// TIA Portal project "GzyHzy_1500" (V15) (continued)
DATA_BLOCK "模拟量"   // DB2
{ S7_Optimized_Access := 'FALSE' }
VERSION : 0.1
   VAR
      STAT0 : Int;
      STAT1 : Int;
      STAT2 : Int;
      STAT3 : Int;
      STAT4 : Int;
      STAT5 : Int;
      STAT6 : Int;
      STAT7 : Int;
      STAT8 : Int;
      STAT9 : Real;
      STAT10 : Real;
      STAT11 : Real;
      STAT12 : Real;
      STAT13 : Real;
      STAT14 : Real;
      STAT15 : Real;
      STAT16 : Real;
      STAT17 : Real;
      STAT18 : Real;
      STAT19 : Real;
      STAT20 : Real;
      STAT21 : Real;
      STAT22 : Real;
      STAT23 : Real;
      STAT24 : Real;
      STAT25 : Real;
      STAT26 : Real;
      STAT27 : Real;
      STAT28 : Real;
      STAT29 : Real;
      STAT30 : Real;
      STAT31 : Real;
      STAT32 : Real;
      STAT33 : Real;
      STAT34 : Real;
      STAT35 : Real;
      STAT36 : Real;
      STAT37 : Real;
      STAT38 : Real;
      STAT39 : Real;
      STAT40 : Real;
      STAT41 : Real;
      STAT42 : Real;
      STAT43 : Real;
      STAT44 : Real;
      STAT45 : Real;
      STAT46 : Real;
      STAT47 : Real;
      STAT48 : Real;
      STAT49 : Real;
      STAT50 : Real;
      STAT51 : Real;
      STAT52 : Real;
      STAT53 : Real;
      STAT54 : Real;
      STAT55 : Real;
      STAT56 : Real;
      STAT57 : Real;
      STAT58 : Real;
      STAT59 : Real;
      STAT60 : Real;
      STAT61 : Real;
      STAT62 : Real;
      STAT63 : Real;
      STAT64 : Real;
      STAT65 : Real;
      STAT66 : Real;
      STAT67 : Real;
      STAT68 : Real;
      STAT69 : Real;
      STAT70 : Real;
      STAT71 : Real;
      STAT72 : Real;
      STAT73 : Real;
      STAT74 : Real;
      STAT75 : Real;
      STAT76 : Real;
      STAT77 : Real;
      STAT78 : Real;
      STAT79 : Real;
      STAT80 : Real;
      STAT81 : Real;
   END_VAR
BEGIN
END_DATA_BLOCK

DATA_BLOCK "给煤机班累计DB块"   // DB3
{ S7_Optimized_Access := 'FALSE' }
VERSION : 0.0
// stored: InstanceOfName 累计功能块
"累计功能块"
BEGIN
END_DATA_BLOCK

DATA_BLOCK "给煤机日累计DB块"   // DB4
{ S7_Optimized_Access := 'FALSE' }
VERSION : 0.0
// stored: InstanceOfName 累计功能块
"累计功能块"
BEGIN
END_DATA_BLOCK

DATA_BLOCK "给煤机总累计DB块"   // DB5
{ S7_Optimized_Access := 'FALSE' }
VERSION : 0.0
// stored: InstanceOfName 累计功能块
"累计功能块"
BEGIN
END_DATA_BLOCK

DATA_BLOCK "DB6_皮带秤粘料"   // DB6
{ S7_Optimized_Access := 'FALSE' }
VERSION : 0.1
   VAR
      干燥窑定量给煤机给定反馈差值 : Real;
      干燥窑定量给煤机给定反馈差值绝对值 : Real;
      real3 : Real;
      real4 : Real;
      real5 : Real;
      real6 : Real;
      real7 : Real;
      real8 : Real;
      real9 : Real;
      real10 : Real;
      real11 : Real;
      real12 : Real;
      real13 : Real;
      real14 : Real;
      real15 : Real;
      real16 : Real;
      real17 : Real;
      real18 : Real;
      real19 : Real;
      real20 : Real;
      干燥窑定量给煤机粘料报警 : Bool;
      bool2 : Bool;
      bool3 : Bool;
      bool4 : Bool;
      bool5 : Bool;
      bool6 : Bool;
      bool7 : Bool;
      bool8 : Bool;
      bool9 : Bool;
      bool10 : Bool;
      bool11 : Bool;
      bool12 : Bool;
      bool13 : Bool;
      bool14 : Bool;
      bool15 : Bool;
      bool16 : Bool;
      bool17 : Bool;
      bool18 : Bool;
      bool19 : Bool;
      bool20 : Bool;
      bool21 : Bool;
   END_VAR
BEGIN
END_DATA_BLOCK

DATA_BLOCK "累计功能块2_DB"   // DB7
{ S7_Optimized_Access := 'FALSE' }
VERSION : 0.1
// stored: InstanceOfName 累计功能块2
"累计功能块2"
BEGIN
END_DATA_BLOCK

DATA_BLOCK "通讯仪表数据"   // DB20
{ S7_Optimized_Access := 'FALSE' }
VERSION : 0.1
   VAR
      STAT0 : Int;
      "1#窑A档油温1" : Real := 33.4;
      "1#窑A档油温2" : Real := 33.0;
      "1#窑A档油温3" : Real := 34.3;
      "1#窑A档油温4" : Real := 34.0;
      "1#窑A档轴温1" : Real := 33.6;
      "1#窑A档轴温2" : Real := 33.4;
      "1#窑A档轴温3" : Real := 33.6;
      "1#窑A档轴温4" : Real := 34.5;
      "1#窑B档油温1" : Real := 34.3;
      "1#窑B档油温2" : Real := 34.5;
      "1#窑B档油温3" : Real := 35.0;
      "1#窑B档油温4" : Real := 36.1;
      "1#窑B档轴温1" : Real := 34.9;
      "1#窑B档轴温2" : Real := 36.4;
      "1#窑B档轴温3" : Real := 34.9;
      "1#窑B档轴温4" : Real := 36.2;
      "1#窑主电机A相绕组温度" : Real := 62.7;
      "1#窑主电机B相绕组温度" : Real := 63.4;
      "1#窑主电机C相绕组温度" : Real := 62.0;
      "1#窑主电机前轴承温度" : Real := 45.0;
      "1#窑主电机后轴承温度" : Real := 41.8;
      STAT22 : Real;
      STAT23 : Real;
      STAT24 : Real;
      STAT25 : Real;
      STAT26 : Real;
      STAT27 : Real;
      STAT28 : Real;
      STAT29 : Real;
      STAT30 : Real;
      STAT31 : Real;
      STAT32 : Real;
      "1#干燥窑煤粉仓称重" : Real := 11.52;   // 1#干燥窑煤粉仓称重
      STAT34 : Real;
   END_VAR
BEGIN
END_DATA_BLOCK

DATA_BLOCK "模拟量数据"   // DB21
{ S7_Optimized_Access := 'FALSE' }
VERSION : 0.1
   VAR
      "1#干燥窑主电机转速" : Real := 795.8328;
      "1#干燥窑主电机电流" : Real := 246.3866;
      STAT2 : Real;
      "1#干燥窑一次风机运行电流" : Real := 48.19213;
      "1#二次风机运行频率" : Real := 29.89005;
      "1#二次风机运行电流" : Real := 89.02026;
      "1#干燥窑窑尾烟气管道压力" : Real := -16.14584;
      "1#备用一次风机运行电流" : Real := 48.94907;
      "1#备用二次风机运行频率" : Real := 0.1157407;
      "1#备用二次风机运行电流" : Real;
      "1#干燥窑煤粉流量" : Real := 2.039641;
      "1#干燥窑进口烟气管道压力" : Real := -66.84027;
      "1#干燥窑一次风机压力" : Real := 2421.875;
      "1#干燥窑二次风机压力" : Real := 1265.625;
      "1#干燥窑煤粉仓压力" : Real := 11.63208;
      "1#干燥窑燃烧室压力" : Real := -751.3021;
      "1#干燥窑煤粉仓温度1" : Real := 17.85301;
      "1#干燥窑煤粉仓温度2" : Real := 35.30093;
      "1#干燥窑煤粉仓温度3" : Real := 33.96991;
      "1#干燥窑煤粉仓温度4" : Real := 35.3588;
      "1#干燥窑窑尾罩温度" : Real := 194.8495;
      "1#干燥窑进口烟气管道温度" : Real := 346.0648;
      "1#干燥窑燃烧室温度" : Real := 883.3333;
      "1#干燥窑混合室温度" : Real := 426.1863;
      "1#干燥窑主机转速给定" : Real := 800.0;
      "1#干燥窑煤粉仓流量给定" : Real := 2.0;
      振动筛转速给定 : Real;
      STAT27 : Real;
      STAT28 : Real;
      "1#二次风机频率给定" : Real := 30.0;
      STAT30 : Real;
      "1#备用二次风机频率给定" : Real := 38.0;
      "1#干燥窑定量给煤机班累计" : Real := 0.004813849;
      "1#干燥窑定量给煤机日累计" : Real := 362.4617;
      "1#干燥窑定量给煤机总累计" : Real := 362.4611;
      STAT35 : Real;
      STAT36 : Real;
      振动筛转速 : Real;
      振动筛电流 : Real;
   END_VAR
BEGIN
END_DATA_BLOCK

DATA_BLOCK "窑联锁"   // DB23
{ S7_Optimized_Access := 'FALSE' }
VERSION : 0.1
   VAR
      STAT0 : Bool := TRUE;
      STAT1 : Bool;
      STAT2 : Bool;
      STAT3 : Bool;
      STAT4 : Bool;
      STAT5 : Bool;
      STAT6 : Bool;
      STAT7 : Bool;
      STAT8 : Bool := TRUE;
      STAT9 : Bool;
      STAT10 : Bool;
      STAT11 : Bool;
      STAT12 : Bool;
      STAT13 : Bool;
      STAT14 : Bool;
      STAT15 : Bool;
      STAT16 : Bool;
      STAT17 : Bool;
      STAT18 : Word;
   END_VAR
BEGIN
END_DATA_BLOCK

DATA_BLOCK "DB26"   // DB26
{ S7_Optimized_Access := 'FALSE' }
VERSION : 0.1
   VAR
      STAT0 : Bool;
      STAT1 : Bool;
      STAT2 : Bool;
      STAT3 : Bool;
      STAT4 : Bool;
      STAT5 : Bool;
      STAT6 : Bool;
      STAT7 : Bool;
      STAT8 : Word := WORD#16#0002;
      STAT9 : Word;
      STAT10 : Word;
   END_VAR
BEGIN
END_DATA_BLOCK

DATA_BLOCK "FB40_DATA_ALARM_DB"   // DB40
{ S7_Optimized_Access := 'FALSE' }
VERSION : 0.1
// stored: InstanceOfName FB40_DATA_ALARM
"FB40_DATA_ALARM"
BEGIN
END_DATA_BLOCK

FUNCTION_BLOCK "累计功能块"   // FB10, STL
{ S7_Optimized_Access := 'FALSE' }
VERSION : 0.1
   VAR_INPUT
      IN0 : Real;
      IN1 : Bool;
   END_VAR
   VAR_OUTPUT
      OUT2 : Real;
   END_VAR
   VAR
      STAT3 : Real;
      STAT4 : Real;
      STAT5 : Real;
   END_VAR
BEGIN

REGION Network 1
         A(;
         A(;
         A(;
         L     #IN0;
         L     3600.0;
         /R;
         T     #STAT3;
         AN    OV;
         SAVE;
         CLR;
         A     BR;
         );
         JNB   M001;
         L     #STAT3;
         L     10.0;
         /R;
         T     #STAT4;
         AN    OV;
         SAVE;
         CLR;
   M001: A     BR;
         );
         JNB   M002;
         L     #STAT4;
         L     #STAT5;
         +R;
         T     #STAT5;
         AN    OV;
         SAVE;
         CLR;
   M002: A     BR;
         );
         JNB   M003;
         L     #STAT5;
         T     #OUT2;
   M003: NOP   0;
END_REGION

REGION Network 2
         A     #IN1;
         =     %L0.0;
         A     %L0.0;
         JNB   M004;
         L     0.0;
         T     #STAT3;
   M004: NOP   0;
         A     %L0.0;
         JNB   M005;
         L     0.0;
         T     #STAT4;
   M005: NOP   0;
         A     %L0.0;
         JNB   M006;
         L     0.0;
         T     #STAT5;
   M006: NOP   0;
END_REGION

REGION Network 3
         SET;
         SAVE;
END_REGION
END_FUNCTION_BLOCK

FUNCTION_BLOCK "FB40_DATA_ALARM"   // FB40, LAD
{ S7_Optimized_Access := 'FALSE' }
VERSION : 0.1
   VAR
      "1#干燥窑主传动转速" : "FB330_DATA_ALARM";
      "1#干燥窑主传动电流" : "FB330_DATA_ALARM";
      "1#干燥窑二次风机电流" : "FB330_DATA_ALARM";
      "1#干燥窑一次风机电流" : "FB330_DATA_ALARM";
      "1#干燥窑二次风机频率" : "FB330_DATA_ALARM";
      "1#干燥窑窑尾压力" : "FB330_DATA_ALARM";
      "1#干燥窑备用一次风机频率" : "FB330_DATA_ALARM";
      "1#干燥窑备用一次风机电流" : "FB330_DATA_ALARM";
      "1#干燥窑备用二次风机频率" : "FB330_DATA_ALARM";
      "1#干燥窑备用二次风机电流" : "FB330_DATA_ALARM";
      定量给煤机流量 : "FB330_DATA_ALARM";
      烟气管道进口压力 : "FB330_DATA_ALARM";
      "1#干燥窑一次风压" : "FB330_DATA_ALARM";
      "1#干燥窑二次风压" : "FB330_DATA_ALARM";
      煤粉仓压力 : "FB330_DATA_ALARM";
      混合室压力 : "FB330_DATA_ALARM";
      "煤粉仓温度1(PT100)" : "FB330_DATA_ALARM";
      "煤粉仓温度2(PT100)" : "FB330_DATA_ALARM";
      "煤粉仓温度3(PT100)" : "FB330_DATA_ALARM";
      "煤粉仓温度4(PT100)" : "FB330_DATA_ALARM";
      "窑尾温度 K偶" : "FB330_DATA_ALARM";
      "烟气管道进口温度 K偶" : "FB330_DATA_ALARM";
      "燃烧室温度 4~20mA" : "FB330_DATA_ALARM";
      "混合室温度 4~20mA" : "FB330_DATA_ALARM";
      "1#干燥窑进料口压力" : "FB330_DATA_ALARM";
      "1#给煤机出料口负压" : "FB330_DATA_ALARM";
      振动筛转速 : "FB330_DATA_ALARM";
      振动筛电流 : "FB330_DATA_ALARM";
      PIW312 : "FB330_DATA_ALARM";
      PIW314 : "FB330_DATA_ALARM";
      PIW316 : "FB330_DATA_ALARM";
      PIW318 : "FB330_DATA_ALARM";
      "1#窑A档轴温1" : "FB330_DATA_ALARM";
      "1#窑A档油温1" : "FB330_DATA_ALARM";
      "1#窑A档轴温2" : "FB330_DATA_ALARM";
      "1#窑A档油温2" : "FB330_DATA_ALARM";
      "1#窑A档轴温3" : "FB330_DATA_ALARM";
      "1#窑A档油温3" : "FB330_DATA_ALARM";
      "1#窑A档轴温4" : "FB330_DATA_ALARM";
      "1#窑A档油温4" : "FB330_DATA_ALARM";
      "1#窑B档轴温1" : "FB330_DATA_ALARM";
      "1#窑B档油温1" : "FB330_DATA_ALARM";
      "1#窑B档轴温2" : "FB330_DATA_ALARM";
      "1#窑B档油温2" : "FB330_DATA_ALARM";
      "1#窑B档轴温3" : "FB330_DATA_ALARM";
      "1#窑B档油温3" : "FB330_DATA_ALARM";
      "1#窑B档轴温4" : "FB330_DATA_ALARM";
      "1#窑B档油温4" : "FB330_DATA_ALARM";
      "1#窑主电机A相绕组温度" : "FB330_DATA_ALARM";
      "1#窑主电机B相绕组温度" : "FB330_DATA_ALARM";
      "1#窑主电机C相绕组温度" : "FB330_DATA_ALARM";
      "1#窑主电机前轴承温度" : "FB330_DATA_ALARM";
      "1#窑主电机后轴承温度" : "FB330_DATA_ALARM";
      PID404 : "FB330_DATA_ALARM";
      PID408 : "FB330_DATA_ALARM";
      PID412 : "FB330_DATA_ALARM";
      "1#干燥窑煤粉仓称重" : "FB330_DATA_ALARM";
      STATIC1 : "FB330_DATA_ALARM";
      STATIC2 : "FB330_DATA_ALARM";
      STATIC3 : "FB330_DATA_ALARM";
   END_VAR
   VAR_TEMP
      TEMP1 : Real;
   END_VAR
BEGIN

REGION Network 1
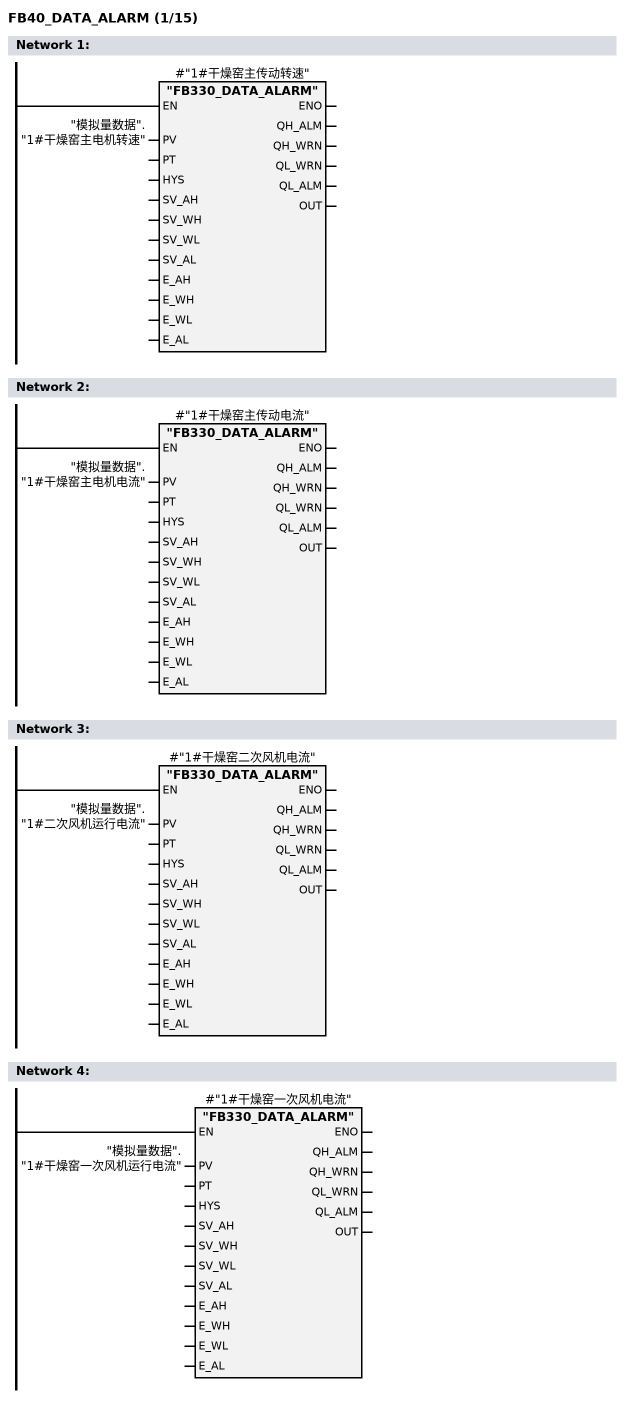
   RUNG wire#powerrail
      #"1#干燥窑主传动转速"(PV := "模拟量数据"."1#干燥窑主电机转速", PT :=, HYS :=, SV_AH :=, SV_WH :=, SV_WL :=, SV_AL :=, E_AH :=, E_WH :=, E_WL :=, E_AL :=, QH_ALM =>, QH_WRN =>, QL_WRN =>, QL_ALM =>, OUT =>)
   END_RUNG
   // the same network as SCL:
   #"1#干燥窑主传动转速"(PV := "模拟量数据"."1#干燥窑主电机转速");   // "FB330_DATA_ALARM"
END_REGION

REGION Network 2
   RUNG wire#powerrail
      #"1#干燥窑主传动电流"(PV := "模拟量数据"."1#干燥窑主电机电流", PT :=, HYS :=, SV_AH :=, SV_WH :=, SV_WL :=, SV_AL :=, E_AH :=, E_WH :=, E_WL :=, E_AL :=, QH_ALM =>, QH_WRN =>, QL_WRN =>, QL_ALM =>, OUT =>)
   END_RUNG
   // the same network as SCL:
   #"1#干燥窑主传动电流"(PV := "模拟量数据"."1#干燥窑主电机电流");   // "FB330_DATA_ALARM"
END_REGION

REGION Network 3
   RUNG wire#powerrail
      #"1#干燥窑二次风机电流"(PV := "模拟量数据"."1#二次风机运行电流", PT :=, HYS :=, SV_AH :=, SV_WH :=, SV_WL :=, SV_AL :=, E_AH :=, E_WH :=, E_WL :=, E_AL :=, QH_ALM =>, QH_WRN =>, QL_WRN =>, QL_ALM =>, OUT =>)
   END_RUNG
   // the same network as SCL:
   #"1#干燥窑二次风机电流"(PV := "模拟量数据"."1#二次风机运行电流");   // "FB330_DATA_ALARM"
END_REGION

REGION Network 4
   RUNG wire#powerrail
      #"1#干燥窑一次风机电流"(PV := "模拟量数据"."1#干燥窑一次风机运行电流", PT :=, HYS :=, SV_AH :=, SV_WH :=, SV_WL :=, SV_AL :=, E_AH :=, E_WH :=, E_WL :=, E_AL :=, QH_ALM =>, QH_WRN =>, QL_WRN =>, QL_ALM =>, OUT =>)
   END_RUNG
   // the same network as SCL:
   #"1#干燥窑一次风机电流"(PV := "模拟量数据"."1#干燥窑一次风机运行电流");   // "FB330_DATA_ALARM"
END_REGION

REGION Network 5
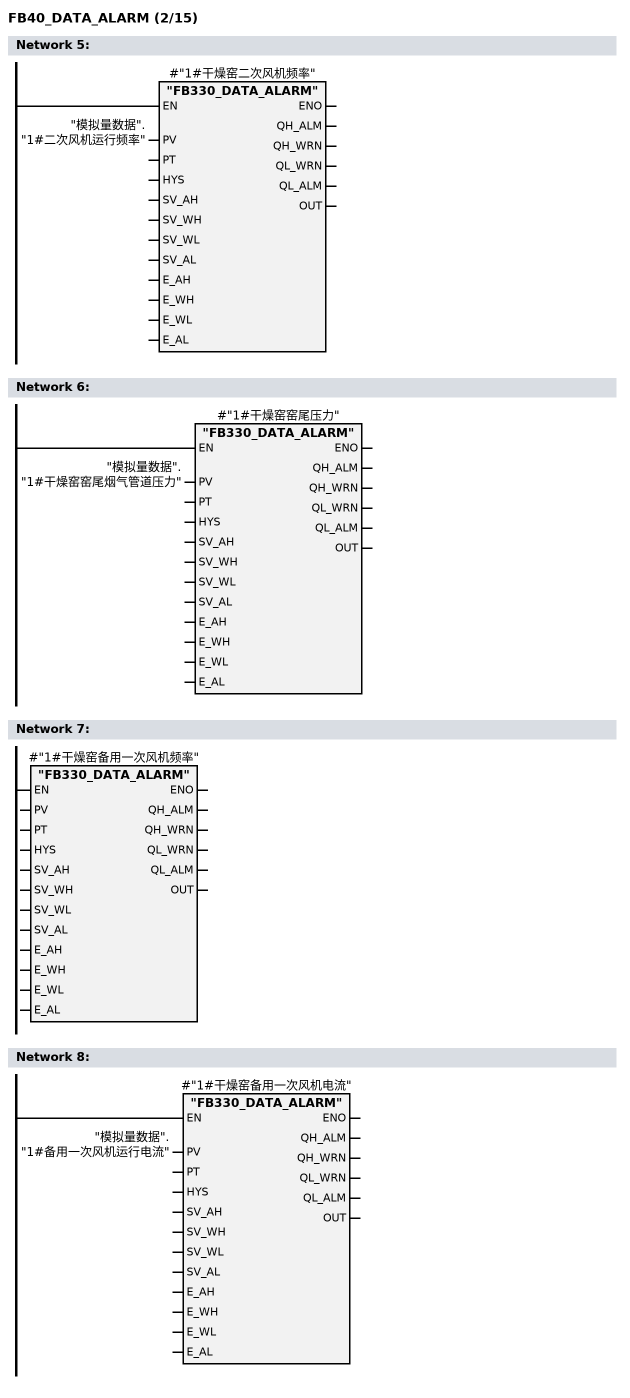
   RUNG wire#powerrail
      #"1#干燥窑二次风机频率"(PV := "模拟量数据"."1#二次风机运行频率", PT :=, HYS :=, SV_AH :=, SV_WH :=, SV_WL :=, SV_AL :=, E_AH :=, E_WH :=, E_WL :=, E_AL :=, QH_ALM =>, QH_WRN =>, QL_WRN =>, QL_ALM =>, OUT =>)
   END_RUNG
   // the same network as SCL:
   #"1#干燥窑二次风机频率"(PV := "模拟量数据"."1#二次风机运行频率");   // "FB330_DATA_ALARM"
END_REGION

REGION Network 6
   RUNG wire#powerrail
      #"1#干燥窑窑尾压力"(PV := "模拟量数据"."1#干燥窑窑尾烟气管道压力", PT :=, HYS :=, SV_AH :=, SV_WH :=, SV_WL :=, SV_AL :=, E_AH :=, E_WH :=, E_WL :=, E_AL :=, QH_ALM =>, QH_WRN =>, QL_WRN =>, QL_ALM =>, OUT =>)
   END_RUNG
   // the same network as SCL:
   #"1#干燥窑窑尾压力"(PV := "模拟量数据"."1#干燥窑窑尾烟气管道压力");   // "FB330_DATA_ALARM"
END_REGION

REGION Network 7
   RUNG wire#powerrail
      #"1#干燥窑备用一次风机频率"(PV :=, PT :=, HYS :=, SV_AH :=, SV_WH :=, SV_WL :=, SV_AL :=, E_AH :=, E_WH :=, E_WL :=, E_AL :=, QH_ALM =>, QH_WRN =>, QL_WRN =>, QL_ALM =>, OUT =>)
   END_RUNG
   // the same network as SCL:
   #"1#干燥窑备用一次风机频率"();   // "FB330_DATA_ALARM"
END_REGION

REGION Network 8
   RUNG wire#powerrail
      #"1#干燥窑备用一次风机电流"(PV := "模拟量数据"."1#备用一次风机运行电流", PT :=, HYS :=, SV_AH :=, SV_WH :=, SV_WL :=, SV_AL :=, E_AH :=, E_WH :=, E_WL :=, E_AL :=, QH_ALM =>, QH_WRN =>, QL_WRN =>, QL_ALM =>, OUT =>)
   END_RUNG
   // the same network as SCL:
   #"1#干燥窑备用一次风机电流"(PV := "模拟量数据"."1#备用一次风机运行电流");   // "FB330_DATA_ALARM"
END_REGION

REGION Network 9
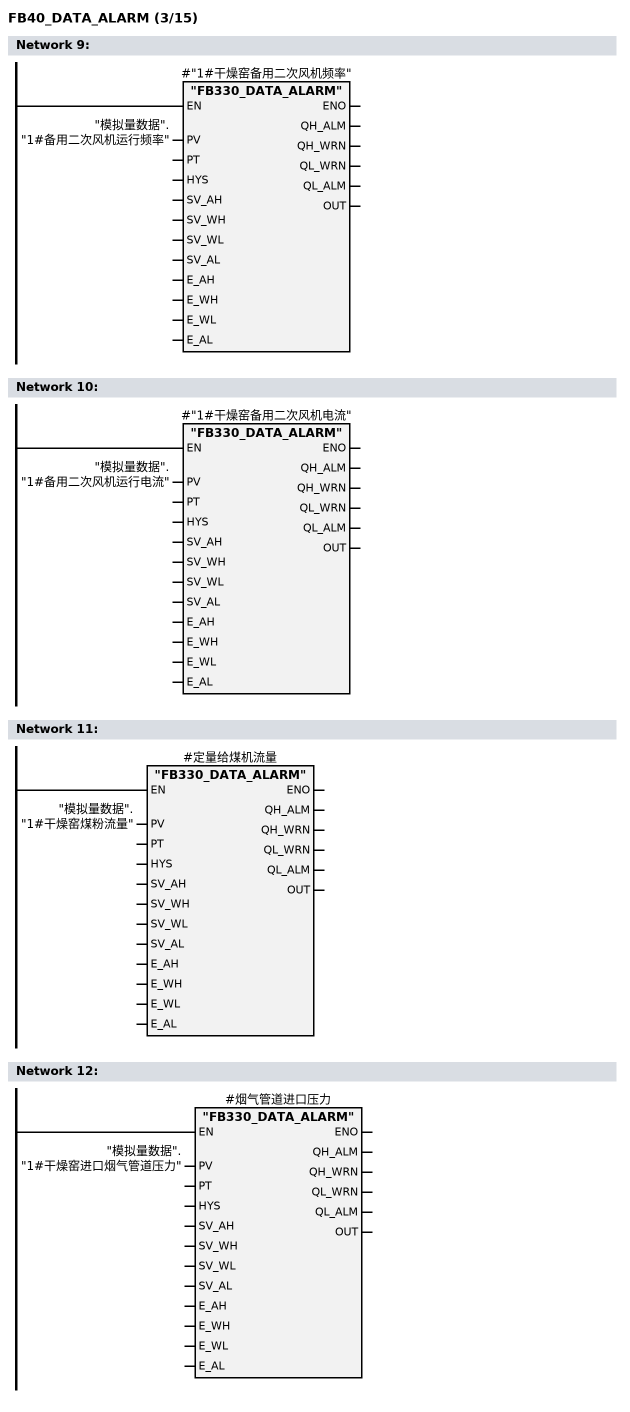
   RUNG wire#powerrail
      #"1#干燥窑备用二次风机频率"(PV := "模拟量数据"."1#备用二次风机运行频率", PT :=, HYS :=, SV_AH :=, SV_WH :=, SV_WL :=, SV_AL :=, E_AH :=, E_WH :=, E_WL :=, E_AL :=, QH_ALM =>, QH_WRN =>, QL_WRN =>, QL_ALM =>, OUT =>)
   END_RUNG
   // the same network as SCL:
   #"1#干燥窑备用二次风机频率"(PV := "模拟量数据"."1#备用二次风机运行频率");   // "FB330_DATA_ALARM"
END_REGION

REGION Network 10
   RUNG wire#powerrail
      #"1#干燥窑备用二次风机电流"(PV := "模拟量数据"."1#备用二次风机运行电流", PT :=, HYS :=, SV_AH :=, SV_WH :=, SV_WL :=, SV_AL :=, E_AH :=, E_WH :=, E_WL :=, E_AL :=, QH_ALM =>, QH_WRN =>, QL_WRN =>, QL_ALM =>, OUT =>)
   END_RUNG
   // the same network as SCL:
   #"1#干燥窑备用二次风机电流"(PV := "模拟量数据"."1#备用二次风机运行电流");   // "FB330_DATA_ALARM"
END_REGION

REGION Network 11
   RUNG wire#powerrail
      #定量给煤机流量(PV := "模拟量数据"."1#干燥窑煤粉流量", PT :=, HYS :=, SV_AH :=, SV_WH :=, SV_WL :=, SV_AL :=, E_AH :=, E_WH :=, E_WL :=, E_AL :=, QH_ALM =>, QH_WRN =>, QL_WRN =>, QL_ALM =>, OUT =>)
   END_RUNG
   // the same network as SCL:
   #定量给煤机流量(PV := "模拟量数据"."1#干燥窑煤粉流量");   // "FB330_DATA_ALARM"
END_REGION

REGION Network 12
   RUNG wire#powerrail
      #烟气管道进口压力(PV := "模拟量数据"."1#干燥窑进口烟气管道压力", PT :=, HYS :=, SV_AH :=, SV_WH :=, SV_WL :=, SV_AL :=, E_AH :=, E_WH :=, E_WL :=, E_AL :=, QH_ALM =>, QH_WRN =>, QL_WRN =>, QL_ALM =>, OUT =>)
   END_RUNG
   // the same network as SCL:
   #烟气管道进口压力(PV := "模拟量数据"."1#干燥窑进口烟气管道压力");   // "FB330_DATA_ALARM"
END_REGION

REGION Network 13
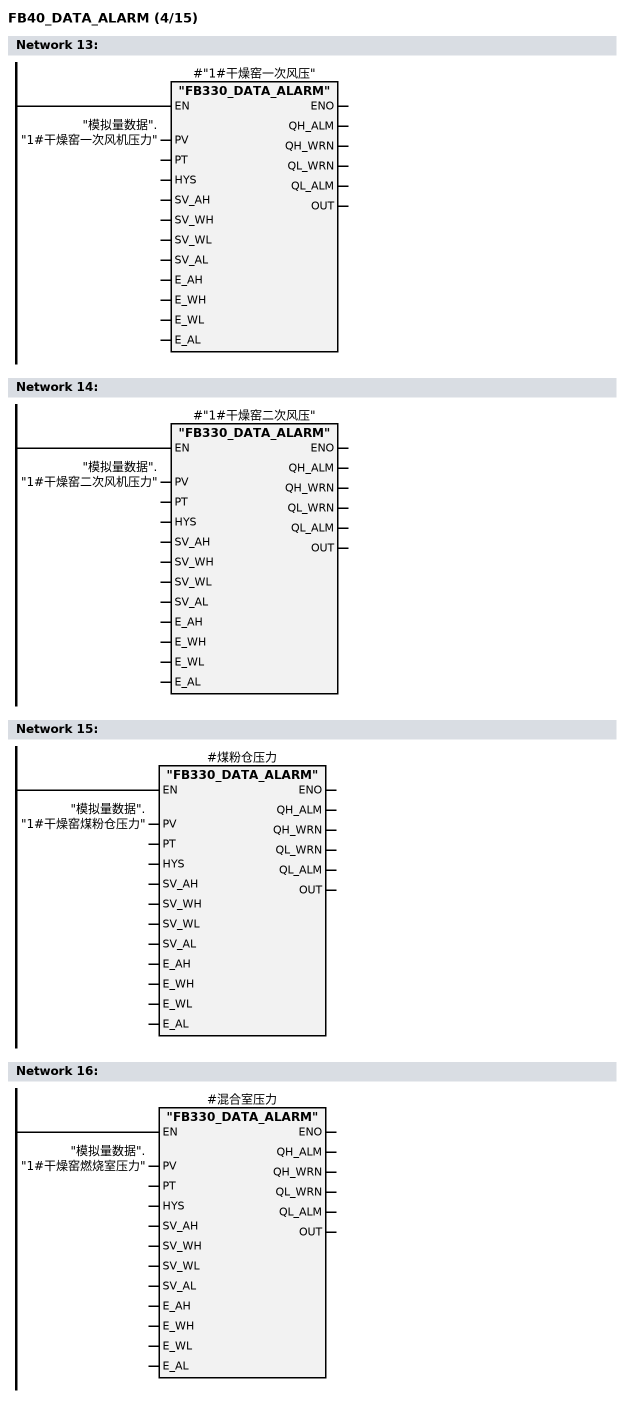
   RUNG wire#powerrail
      #"1#干燥窑一次风压"(PV := "模拟量数据"."1#干燥窑一次风机压力", PT :=, HYS :=, SV_AH :=, SV_WH :=, SV_WL :=, SV_AL :=, E_AH :=, E_WH :=, E_WL :=, E_AL :=, QH_ALM =>, QH_WRN =>, QL_WRN =>, QL_ALM =>, OUT =>)
   END_RUNG
   // the same network as SCL:
   #"1#干燥窑一次风压"(PV := "模拟量数据"."1#干燥窑一次风机压力");   // "FB330_DATA_ALARM"
END_REGION

REGION Network 14
   RUNG wire#powerrail
      #"1#干燥窑二次风压"(PV := "模拟量数据"."1#干燥窑二次风机压力", PT :=, HYS :=, SV_AH :=, SV_WH :=, SV_WL :=, SV_AL :=, E_AH :=, E_WH :=, E_WL :=, E_AL :=, QH_ALM =>, QH_WRN =>, QL_WRN =>, QL_ALM =>, OUT =>)
   END_RUNG
   // the same network as SCL:
   #"1#干燥窑二次风压"(PV := "模拟量数据"."1#干燥窑二次风机压力");   // "FB330_DATA_ALARM"
END_REGION

REGION Network 15
   RUNG wire#powerrail
      #煤粉仓压力(PV := "模拟量数据"."1#干燥窑煤粉仓压力", PT :=, HYS :=, SV_AH :=, SV_WH :=, SV_WL :=, SV_AL :=, E_AH :=, E_WH :=, E_WL :=, E_AL :=, QH_ALM =>, QH_WRN =>, QL_WRN =>, QL_ALM =>, OUT =>)
   END_RUNG
   // the same network as SCL:
   #煤粉仓压力(PV := "模拟量数据"."1#干燥窑煤粉仓压力");   // "FB330_DATA_ALARM"
END_REGION

REGION Network 16
   RUNG wire#powerrail
      #混合室压力(PV := "模拟量数据"."1#干燥窑燃烧室压力", PT :=, HYS :=, SV_AH :=, SV_WH :=, SV_WL :=, SV_AL :=, E_AH :=, E_WH :=, E_WL :=, E_AL :=, QH_ALM =>, QH_WRN =>, QL_WRN =>, QL_ALM =>, OUT =>)
   END_RUNG
   // the same network as SCL:
   #混合室压力(PV := "模拟量数据"."1#干燥窑燃烧室压力");   // "FB330_DATA_ALARM"
END_REGION

REGION Network 17
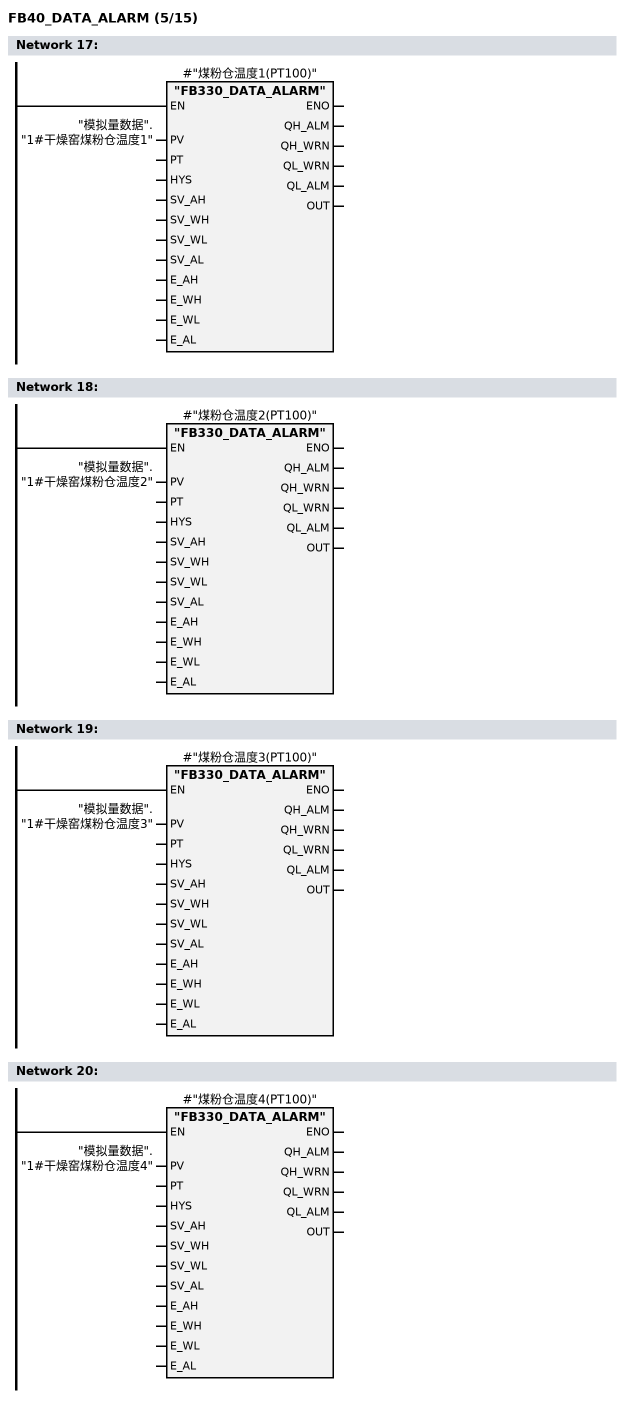
   RUNG wire#powerrail
      #"煤粉仓温度1(PT100)"(PV := "模拟量数据"."1#干燥窑煤粉仓温度1", PT :=, HYS :=, SV_AH :=, SV_WH :=, SV_WL :=, SV_AL :=, E_AH :=, E_WH :=, E_WL :=, E_AL :=, QH_ALM =>, QH_WRN =>, QL_WRN =>, QL_ALM =>, OUT =>)
   END_RUNG
   // the same network as SCL:
   #"煤粉仓温度1(PT100)"(PV := "模拟量数据"."1#干燥窑煤粉仓温度1");   // "FB330_DATA_ALARM"
END_REGION

REGION Network 18
   RUNG wire#powerrail
      #"煤粉仓温度2(PT100)"(PV := "模拟量数据"."1#干燥窑煤粉仓温度2", PT :=, HYS :=, SV_AH :=, SV_WH :=, SV_WL :=, SV_AL :=, E_AH :=, E_WH :=, E_WL :=, E_AL :=, QH_ALM =>, QH_WRN =>, QL_WRN =>, QL_ALM =>, OUT =>)
   END_RUNG
   // the same network as SCL:
   #"煤粉仓温度2(PT100)"(PV := "模拟量数据"."1#干燥窑煤粉仓温度2");   // "FB330_DATA_ALARM"
END_REGION

REGION Network 19
   RUNG wire#powerrail
      #"煤粉仓温度3(PT100)"(PV := "模拟量数据"."1#干燥窑煤粉仓温度3", PT :=, HYS :=, SV_AH :=, SV_WH :=, SV_WL :=, SV_AL :=, E_AH :=, E_WH :=, E_WL :=, E_AL :=, QH_ALM =>, QH_WRN =>, QL_WRN =>, QL_ALM =>, OUT =>)
   END_RUNG
   // the same network as SCL:
   #"煤粉仓温度3(PT100)"(PV := "模拟量数据"."1#干燥窑煤粉仓温度3");   // "FB330_DATA_ALARM"
END_REGION

REGION Network 20
   RUNG wire#powerrail
      #"煤粉仓温度4(PT100)"(PV := "模拟量数据"."1#干燥窑煤粉仓温度4", PT :=, HYS :=, SV_AH :=, SV_WH :=, SV_WL :=, SV_AL :=, E_AH :=, E_WH :=, E_WL :=, E_AL :=, QH_ALM =>, QH_WRN =>, QL_WRN =>, QL_ALM =>, OUT =>)
   END_RUNG
   // the same network as SCL:
   #"煤粉仓温度4(PT100)"(PV := "模拟量数据"."1#干燥窑煤粉仓温度4");   // "FB330_DATA_ALARM"
END_REGION

REGION Network 21
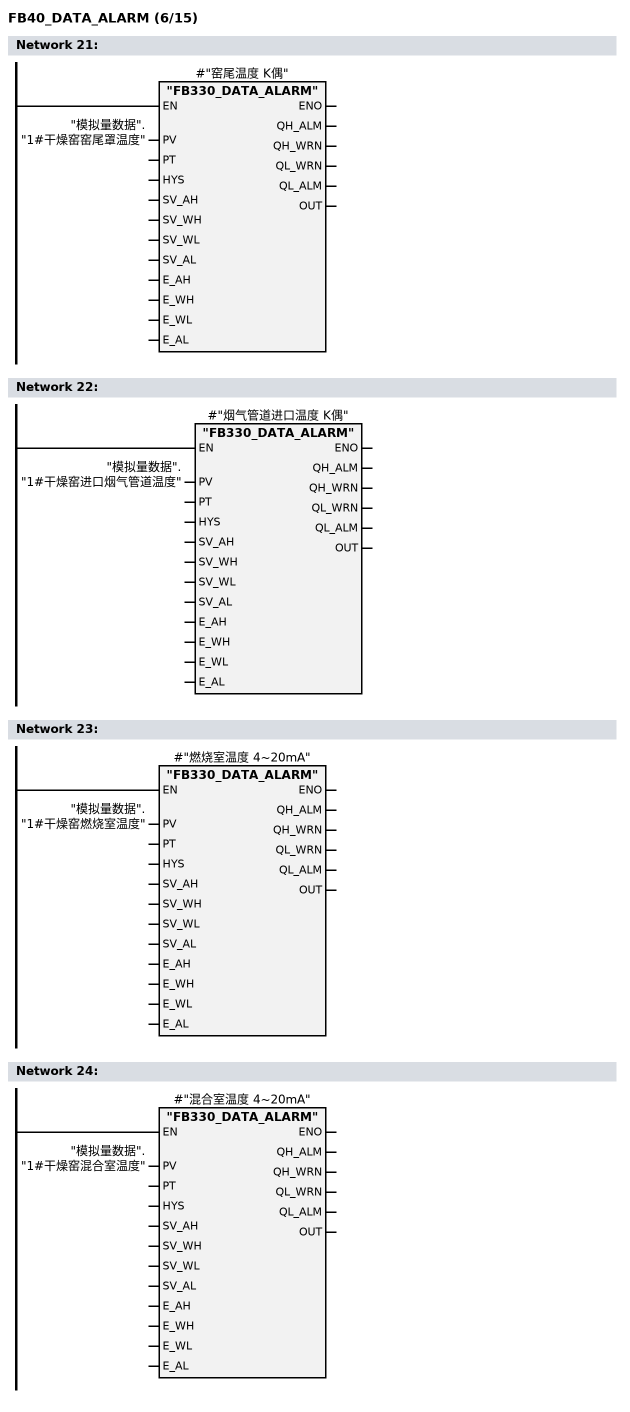
   RUNG wire#powerrail
      #"窑尾温度 K偶"(PV := "模拟量数据"."1#干燥窑窑尾罩温度", PT :=, HYS :=, SV_AH :=, SV_WH :=, SV_WL :=, SV_AL :=, E_AH :=, E_WH :=, E_WL :=, E_AL :=, QH_ALM =>, QH_WRN =>, QL_WRN =>, QL_ALM =>, OUT =>)
   END_RUNG
   // the same network as SCL:
   #"窑尾温度 K偶"(PV := "模拟量数据"."1#干燥窑窑尾罩温度");   // "FB330_DATA_ALARM"
END_REGION

REGION Network 22
   RUNG wire#powerrail
      #"烟气管道进口温度 K偶"(PV := "模拟量数据"."1#干燥窑进口烟气管道温度", PT :=, HYS :=, SV_AH :=, SV_WH :=, SV_WL :=, SV_AL :=, E_AH :=, E_WH :=, E_WL :=, E_AL :=, QH_ALM =>, QH_WRN =>, QL_WRN =>, QL_ALM =>, OUT =>)
   END_RUNG
   // the same network as SCL:
   #"烟气管道进口温度 K偶"(PV := "模拟量数据"."1#干燥窑进口烟气管道温度");   // "FB330_DATA_ALARM"
END_REGION

REGION Network 23
   RUNG wire#powerrail
      #"燃烧室温度 4~20mA"(PV := "模拟量数据"."1#干燥窑燃烧室温度", PT :=, HYS :=, SV_AH :=, SV_WH :=, SV_WL :=, SV_AL :=, E_AH :=, E_WH :=, E_WL :=, E_AL :=, QH_ALM =>, QH_WRN =>, QL_WRN =>, QL_ALM =>, OUT =>)
   END_RUNG
   // the same network as SCL:
   #"燃烧室温度 4~20mA"(PV := "模拟量数据"."1#干燥窑燃烧室温度");   // "FB330_DATA_ALARM"
END_REGION

REGION Network 24
   RUNG wire#powerrail
      #"混合室温度 4~20mA"(PV := "模拟量数据"."1#干燥窑混合室温度", PT :=, HYS :=, SV_AH :=, SV_WH :=, SV_WL :=, SV_AL :=, E_AH :=, E_WH :=, E_WL :=, E_AL :=, QH_ALM =>, QH_WRN =>, QL_WRN =>, QL_ALM =>, OUT =>)
   END_RUNG
   // the same network as SCL:
   #"混合室温度 4~20mA"(PV := "模拟量数据"."1#干燥窑混合室温度");   // "FB330_DATA_ALARM"
END_REGION

REGION Network 25
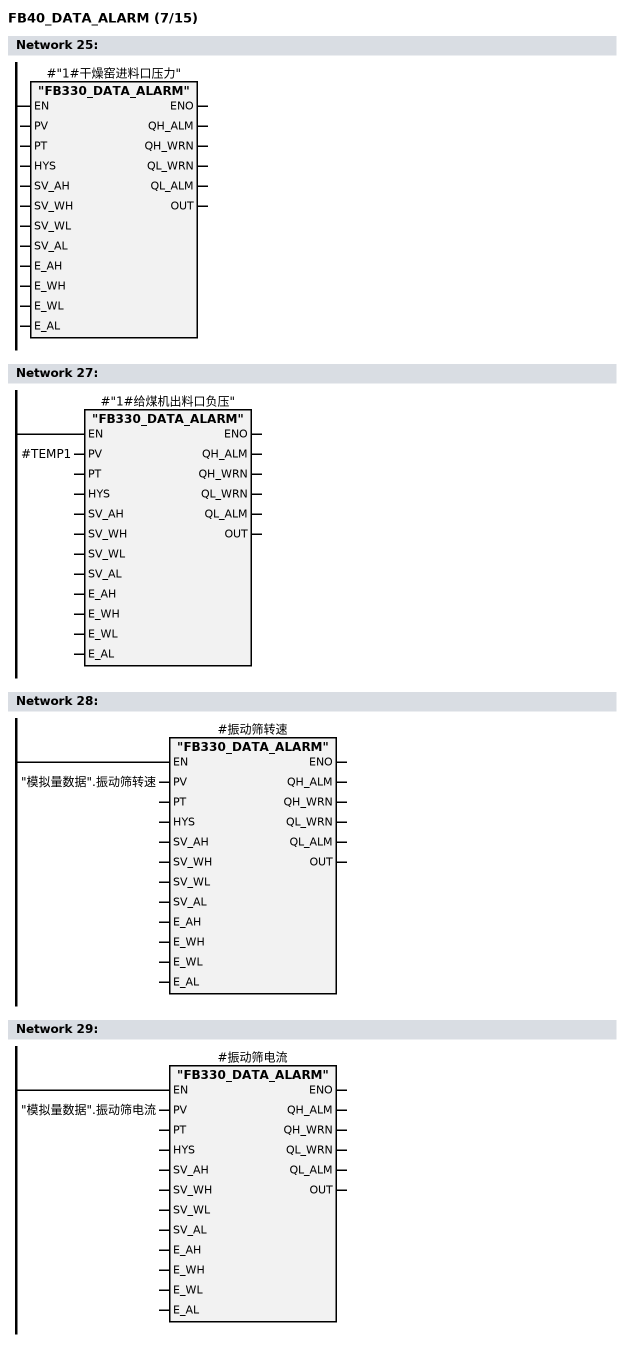
   RUNG wire#powerrail
      #"1#干燥窑进料口压力"(PV :=, PT :=, HYS :=, SV_AH :=, SV_WH :=, SV_WL :=, SV_AL :=, E_AH :=, E_WH :=, E_WL :=, E_AL :=, QH_ALM =>, QH_WRN =>, QL_WRN =>, QL_ALM =>, OUT =>)
   END_RUNG
   // the same network as SCL:
   #"1#干燥窑进料口压力"();   // "FB330_DATA_ALARM"
END_REGION

REGION Network 27
   RUNG wire#powerrail
      #"1#给煤机出料口负压"(PV := #TEMP1, PT :=, HYS :=, SV_AH :=, SV_WH :=, SV_WL :=, SV_AL :=, E_AH :=, E_WH :=, E_WL :=, E_AL :=, QH_ALM =>, QH_WRN =>, QL_WRN =>, QL_ALM =>, OUT =>)
   END_RUNG
   // the same network as SCL:
   #"1#给煤机出料口负压"(PV := #TEMP1);   // "FB330_DATA_ALARM"
END_REGION

REGION Network 28
   RUNG wire#powerrail
      #振动筛转速(PV := "模拟量数据".振动筛转速, PT :=, HYS :=, SV_AH :=, SV_WH :=, SV_WL :=, SV_AL :=, E_AH :=, E_WH :=, E_WL :=, E_AL :=, QH_ALM =>, QH_WRN =>, QL_WRN =>, QL_ALM =>, OUT =>)
   END_RUNG
   // the same network as SCL:
   #振动筛转速(PV := "模拟量数据".振动筛转速);   // "FB330_DATA_ALARM"
END_REGION

REGION Network 29
   RUNG wire#powerrail
      #振动筛电流(PV := "模拟量数据".振动筛电流, PT :=, HYS :=, SV_AH :=, SV_WH :=, SV_WL :=, SV_AL :=, E_AH :=, E_WH :=, E_WL :=, E_AL :=, QH_ALM =>, QH_WRN =>, QL_WRN =>, QL_ALM =>, OUT =>)
   END_RUNG
   // the same network as SCL:
   #振动筛电流(PV := "模拟量数据".振动筛电流);   // "FB330_DATA_ALARM"
END_REGION

REGION Network 30